VERSION : 0.1
   VAR_INPUT
      null_value : DInt;   // value that indicates null data
   END_VAR
   VAR_IN_OUT
      int_array : Variant;
   END_VAR
   VAR_TEMP
      i : Int;
      j : Int;
      len_int : Int;
      len_udint : UDInt;
      status : Int;
      t_int_array : Array[0..999] of DInt;
   END_VAR
BEGIN
   REGION "COPY TO LOCAL MEMORY"
       #len_udint := CountOfElements(#int_array);
       #len_int := UDINT_TO_INT(#len_udint) - 1;
       #status := MOVE_BLK_VARIANT(SRC := #int_array,
                                   COUNT := #len_udint,
                                   SRC_INDEX := 0,
                                   DEST_INDEX := 0,
                                   DEST => #t_int_array);
   END_REGION

   REGION "COLLAPSE IN PLACE"
       FOR #i := 0 TO #len_int - 1 DO
           IF #t_int_array[#i] = #null_value THEN
               FOR #j := #i + 1 TO #len_int DO
                   IF #t_int_array[#j] <> #null_value THEN
                       #t_int_array[#i] := #t_int_array[#j];
                       #t_int_array[#j] := #null_value;
                       EXIT;
                   END_IF;
               END_FOR;
           END_IF;
       END_FOR;
   END_REGION

   REGION "RETURN"
       #status := MOVE_BLK_VARIANT(SRC := #t_int_array,
                                   COUNT := #len_udint,
                                   SRC_INDEX := 0,
                                   DEST_INDEX := 0,
                                   DEST => #int_array);
   END_REGION
END_FUNCTION

FUNCTION "Count Collapsed DInt Array" : Int   // FC133, SCL
{ S7_Optimized_Access := 'TRUE' }
VERSION : 0.1
   VAR_INPUT
      null_value : DInt;
      "array" : Variant;
   END_VAR
   VAR_TEMP
      count : Int;
      i : Int;
      len_int : Int;
      len_udint : UDInt;
      status : Int;
      t_array : Array[0..999] of DInt;
   END_VAR
BEGIN
   REGION "NOTES"
       (*
       returns the number of valid elements in a collapsed int array
       *)
   END_REGION


   REGION "COPY TO LOCAL"
       #len_udint := CountOfElements(#array);
       #len_int := UDINT_TO_INT(#len_udint) - 1;
       #status := MOVE_BLK_VARIANT(SRC := #array,
                                   COUNT := #len_udint,
                                   SRC_INDEX := 0,
                                   DEST_INDEX := 0,
                                   DEST => #t_array);
   END_REGION


   REGION "SCAN FOR FIRST NULL"
       FOR #i := 0 TO #len_int DO
           IF #t_array[#i] = INT_TO_DINT("NULL_TOKEN") THEN
               EXIT;
           END_IF;
           IF #t_array[#i] <> #null_value THEN
               #count += 1;
           END_IF;
       END_FOR;
   END_REGION


   REGION "RETURN"
       #"Count Collapsed DInt Array" := #count;
   END_REGION
END_FUNCTION

FUNCTION "Map WIP Codes to DInt Array" : Void   // FC139, SCL
{ S7_Optimized_Access := 'TRUE' }
VERSION : 0.1
   VAR_INPUT
      station : "WIP: Station";
   END_VAR
   VAR_IN_OUT
      WIP_array : Array[0.."WIP_COUNT"] of DInt;
   END_VAR
   VAR_TEMP
      i : Int;
   END_VAR
BEGIN
   FOR #i := 0 TO "WIP_COUNT" DO
       IF #station.wip[#i].wip.code = "NULL_TOKEN" THEN
           EXIT;
       END_IF;
       #WIP_array[#i] := #station.wip[#i].wip.code;
   END_FOR;
END_FUNCTION

FUNCTION "Map Selected Stations to Int Array" : Void   // FC142, SCL
{ S7_Optimized_Access := 'TRUE' }
VERSION : 0.1
   VAR_INPUT
      selected_stations : "Selected Stations";
   END_VAR
   VAR_OUTPUT
      selected_stations_indicies : Array[0.."STATION_COUNT"] of Int;
   END_VAR
   VAR_TEMP
      i : Int;
      p_ret : Int;
      _return : Array[0.."STATION_COUNT"] of Int;
   END_VAR
BEGIN
   "Array.Int.Fill"(value := "NULL_TOKEN",
                    int_array := #_return);
   FOR #i := 0 TO "STATION_COUNT" DO
       IF #selected_stations.stns[#i] THEN
           #_return[#p_ret] := #i;
           #p_ret += 1;
       END_IF;
   END_FOR;
   #selected_stations_indicies := #_return;
END_FUNCTION

FUNCTION "Part_Number_Double.USInt_State_Change" : "State Changes: USInt"   // FC258, SCL
{ S7_Optimized_Access := 'TRUE' }
VERSION : 0.1
   VAR_INPUT
      interface : USInt;
      old : USInt;
   END_VAR
   VAR_TEMP
      _return : "State Changes: USInt";
   END_VAR
BEGIN
       #_return.rising := "USInt.Value_Change"(value := #interface,
                                               old_value := #old);
       #_return.actual := #interface;
       #_return.falling := FALSE;     // animate never set to null token 
       #"Part_Number_Double.USInt_State_Change" := #_return;
END_FUNCTION

FUNCTION "Part_Number_Double.Bool_State_Change" : "State Changes: Bool"   // FC259, SCL
{ S7_Optimized_Access := 'TRUE' }
VERSION : 0.1
   VAR_INPUT
      interface : Bool;
      old : Bool;
   END_VAR
   VAR_TEMP
      _return : "State Changes: Bool";
   END_VAR
BEGIN
   #_return.rising := "Bool.Rising_Edge"(signal := #interface,
                                                 old_signal := #old);
   #_return.actual := #interface;
   #_return.falling := "Bool.Falling_Edge"(signal := #interface,
                                           old_signal := #old);
   #"Part_Number_Double.Bool_State_Change" := #_return;
END_FUNCTION

FUNCTION "Part_Number_Double.WString_State_Change" : "State Changes: WString"   // FC260, SCL
{ S7_Optimized_Access := 'TRUE' }
VERSION : 0.1
   VAR_INPUT
      interface : WString;
      old : WString;
   END_VAR
   VAR_TEMP
      _return : "State Changes: WString";
   END_VAR
BEGIN
   #_return.rising := "WString.Rising_Edge"(value := #interface,
                                             old_value := #old);
   #_return.actual := #interface;
   #_return.falling := "WString.Falling_Edge"(value := #interface,
                                               old_value := #old);
   #"Part_Number_Double.WString_State_Change" := #_return;
END_FUNCTION

FUNCTION "Part_Number_Double_IO_Field.Set_Mode" : Void   // FC261, SCL
{ S7_Optimized_Access := 'TRUE' }
VERSION : 0.1
   VAR_INPUT
      feedback : "Part_Number_Double.State_Change.UDT";
   END_VAR
   VAR_IN_OUT
      mode : String;
   END_VAR
   VAR CONSTANT
      SINGLE : String := 'single';
      DOUBLE : String := 'double';
   END_VAR
BEGIN
   IF #mode = #SINGLE AND #feedback.single.actuate.falling THEN
       #mode := #DOUBLE;
       RETURN;
   END_IF;

   IF #mode = #DOUBLE AND #feedback.double.actuate.falling THEN
       #mode := #SINGLE;
       RETURN;
   END_IF;
END_FUNCTION

FUNCTION "Array.Table_Row.Copy" : Void   // FC296, SCL
{ S7_Optimized_Access := 'TRUE' }
VERSION : 0.1
   VAR_INPUT
      source : Array[*] of "Table Row";
   END_VAR
   VAR_IN_OUT
      destination : Array[*] of "Table Row";
   END_VAR
   VAR_TEMP
      _length_source : DInt;
      _length_destination : DInt;
      _upper_bound : DInt;
      _i : DInt;
   END_VAR
BEGIN
   REGION "FIND UPPER BOUND"
       #_length_source := UDINT_TO_DINT("Array.Any.Length"(#source)) - 1;
       #_length_destination := UDINT_TO_DINT("Array.Any.Length"(#destination)) - 1;
       #_upper_bound := #_length_source;
       IF #_length_destination < #_length_source THEN
           #_upper_bound := #_length_destination;
       END_IF;
   END_REGION


   REGION "PERFORM COPY"
       FOR #_i := 0 TO #_upper_bound DO
           #destination[#_i] := #source[#_i];
       END_FOR;
   END_REGION


   REGION "RETURN"    
       RETURN;
   END_REGION
END_FUNCTION

// folder: Utilities/Address

FUNCTION "Address.Get_Button" : DInt   // FC21, SCL
{ S7_Optimized_Access := 'TRUE' }
VERSION : 0.1
   VAR_INPUT
      address : DInt;
   END_VAR
BEGIN
   #"Address.Get_Button" := #address MOD 10;
END_FUNCTION

FUNCTION "Address.Get_Station" : DInt   // FC24, SCL
{ S7_Optimized_Access := 'TRUE' }
VERSION : 0.1
   VAR_INPUT
      address : DInt;
   END_VAR
BEGIN
   #"Address.Get_Station" := #address / 10_000;
END_FUNCTION

FUNCTION "Address.Set_Address" : DInt   // FC32, SCL
{ S7_Optimized_Access := 'TRUE' }
VERSION : 0.1
   VAR_INPUT
      pBtn : Int;
      pStn : Int;
      pWip : Int;
   END_VAR
BEGIN
   #"Address.Set_Address" := INT_TO_DINT(#pStn) * 10_000 + INT_TO_DINT(#pWip) * 10 + INT_TO_DINT(#pBtn);
END_FUNCTION

FUNCTION "Address.Get_Wip" : DInt   // FC88, SCL
{ S7_Optimized_Access := 'TRUE' }
VERSION : 0.1
   VAR_INPUT
      address : DInt;
   END_VAR
BEGIN
   #"Address.Get_Wip" := #address - "Address.Get_Station"(#address) * 10_000 - "Address.Get_Button"(#address);
END_FUNCTION

// folder: Utilities/Array

FUNCTION "Array.Any.Length" : UDInt   // FC60, SCL
{ S7_Optimized_Access := 'TRUE' }
VERSION : 0.1
   VAR_INPUT
      "array" : Variant;
   END_VAR
   VAR_TEMP
      status : DInt;
      ret : UDInt;
   END_VAR
BEGIN
   #ret := CountOfElements(#array);
   #"Array.Any.Length" := #ret;
END_FUNCTION

FUNCTION "Get Station Index From Id" : Int   // FC106, SCL
{ S7_Optimized_Access := 'TRUE' }
VERSION : 0.1
   VAR_INPUT
      line_name : WString;
      drop_zone : USInt;
      stns : "Station: All Stations";
   END_VAR
   VAR_TEMP
      i : Int;
      ret : Int;
   END_VAR
BEGIN
   REGION "MATCH LINE NAME AND DROP ZONE"
       FOR #i := 0 TO "STATION_COUNT" DO
           IF #line_name = #stns.stn[#i].id.lineName THEN
               IF #drop_zone = #stns.stn[#i].id.dropZone THEN
                   #ret := #i;
                   EXIT;
               END_IF;
           END_IF;
       END_FOR;
   END_REGION


   REGION "RETURN"
       #"Get Station Index From Id" := #ret;
   END_REGION
END_FUNCTION

FUNCTION "Array.Int.Fill" : Void   // FC109, SCL
{ S7_Optimized_Access := 'TRUE' }
VERSION : 0.1
   VAR_INPUT
      value : Int;
   END_VAR
   VAR_IN_OUT
      int_array : Array[*] of Int;
   END_VAR
   VAR_TEMP
      _i : DInt;
      _length : DInt;
   END_VAR
BEGIN
   REGION "GET LENGHT"
       #_length := UDINT_TO_DINT("Array.Any.Length"(#int_array));
       #_length -= 1;
   END_REGION


   REGION "FILL LENGTH WITH BYTE IN"
       FOR #_i := 0 TO #_length DO
           #int_array[#_i] := #value;
       END_FOR;
   END_REGION
END_FUNCTION

FUNCTION "Array.DInt.Is_Element" : Bool   // FC111, SCL
{ S7_Optimized_Access := 'TRUE' }
VERSION : 0.1
   VAR_INPUT
      dint_array : Array[*] of DInt;
      search_term : DInt;
   END_VAR
   VAR_TEMP
      _i : DInt;
      _length : DInt;
   END_VAR
BEGIN
   REGION "LOCAL VARIABLES"
       #_length := UDINT_TO_DINT("Array.Any.Length"(#dint_array)) - 1;
   END_REGION


   REGION "SEARCH ARRAY"
       FOR #_i := 0 TO #_length DO
           IF #dint_array[#_i] <> #search_term THEN
               CONTINUE;
           END_IF;
           #"Array.DInt.Is_Element" := TRUE;
           RETURN;
       END_FOR;
   END_REGION


   REGION "NOT FOUND"
       #"Array.DInt.Is_Element" := FALSE;
       RETURN;
   END_REGION
END_FUNCTION

FUNCTION "Array.Int.Collapse" : Void   // FC114, SCL
{ S7_Optimized_Access := 'TRUE' }
VERSION : 0.1
   VAR_INPUT
      null_value : Int;   // value that indicates null data
   END_VAR
   VAR_IN_OUT
      int_array : Variant;
   END_VAR
   VAR_TEMP
      i : Int;
      j : Int;
      len_int : Int;
      len_udint : UDInt;
      status : Int;
      t_int_array : Array[0..999] of Int;
   END_VAR
BEGIN
   REGION "COPY TO LOCAL MEMORY"
       #len_udint := CountOfElements(#int_array);
       #len_int := UDINT_TO_INT(#len_udint) - 1;
       #status := MOVE_BLK_VARIANT(SRC := #int_array,
                                   COUNT := #len_udint,
                                   SRC_INDEX := 0,
                                   DEST_INDEX := 0,
                                   DEST => #t_int_array);
   END_REGION

   REGION "COLLAPSE IN PLACE"
       FOR #i := 0 TO #len_int - 1 DO
           IF #t_int_array[#i] = #null_value THEN
               FOR #j := #i + 1 TO #len_int DO
                   IF #t_int_array[#j] <> #null_value THEN
                       #t_int_array[#i] := #t_int_array[#j];
                       #t_int_array[#j] := #null_value;
                       EXIT;
                   END_IF;
               END_FOR;
           END_IF;
       END_FOR;
   END_REGION

   REGION "RETURN"
       #status := MOVE_BLK_VARIANT(SRC := #t_int_array,
                                   COUNT := #len_udint,
                                   SRC_INDEX := 0,
                                   DEST_INDEX := 0,
                                   DEST => #int_array);
   END_REGION
END_FUNCTION

FUNCTION "Array.Int.Count" : Int   // FC115, SCL
{ S7_Optimized_Access := 'TRUE' }
VERSION : 0.1
   VAR_INPUT
      null_value : Int;
      "array" : Variant;
   END_VAR
   VAR_TEMP
      count : Int;
      i : Int;
      len_int : Int;
      len_udint : UDInt;
      status : Int;
      t_array : Array[0..999] of Int;
   END_VAR
BEGIN
   REGION "NOTES"
       (*
       returns the number of valid elements in a collapsed int array
       *)
   END_REGION


   REGION "COPY TO LOCAL"
       #len_udint := CountOfElements(#array);
       #len_int := UDINT_TO_INT(#len_udint) - 1;
       #status := MOVE_BLK_VARIANT(SRC := #array,
                                   COUNT := #len_udint,
                                   SRC_INDEX := 0,
                                   DEST_INDEX := 0,
                                   DEST => #t_array);
   END_REGION


   REGION "SCAN FOR FIRST NULL"
       FOR #i := 0 TO #len_int DO
           IF #t_array[#i] = #null_value THEN
               EXIT;
           END_IF;
           IF #t_array[#i] <> #null_value THEN
               #count += 1;
           END_IF;
       END_FOR;
   END_REGION


   REGION "RETURN"
       #"Array.Int.Count" := #count;
   END_REGION
END_FUNCTION

FUNCTION "Array.Bool.True_Indices" : Void   // FC120, SCL
{ S7_Optimized_Access := 'TRUE' }
VERSION : 0.1
   VAR_INPUT
      array_of_bool : Array[*] of Bool;   // max 1000 elements
      length : Int;   // necessary because dynamically sized arrays of bool get passed as arrays with size of a multiple of 8
   END_VAR
   VAR_IN_OUT
      list_of_indices : Array[*] of Int;   // max 1000 elements
   END_VAR
   VAR_TEMP
      _i : Int;
      _p_return : Int;
      _resized_bool_array : Array[0..#UBOUND] of Bool;
   END_VAR
   VAR CONSTANT
      UBOUND : Int := 999;
   END_VAR
BEGIN
   REGION "FILL RETURN ARRAY"
       "Array.Int.Fill"(value := "NULL_TOKEN",
                        int_array := #list_of_indices);
   END_REGION


   REGION "COPY TO ARRAY OF STATIC SIZE"
       FOR #_i := 0 TO #length DO
           #_resized_bool_array[#_i] := #array_of_bool[#_i];
       END_FOR;
   END_REGION


   REGION "INSERT INDICES INTO RETURN ARRAY"
       FOR #_i := 0 TO #length DO
           IF #_resized_bool_array[#_i] THEN
               #list_of_indices[#_p_return] := #_i;
               #_p_return += 1;
           END_IF;
       END_FOR;
   END_REGION
END_FUNCTION

FUNCTION "Array.Int.Is_Element" : Bool   // FC121, SCL
{ S7_Optimized_Access := 'TRUE' }
VERSION : 0.1
   VAR_INPUT
      int_array : Array[*] of Int;
      search_term : Int;
   END_VAR
   VAR_TEMP
      _i : Int;
      _length : DInt;
   END_VAR
BEGIN
   REGION "LOCAL VARIABLES"
       #_length := UDINT_TO_DINT("Array.Any.Length"(#int_array)) - 1;
   END_REGION


   REGION "SEARCH ARRAY"
       FOR #_i := 0 TO #_length DO
           IF #int_array[#_i] <> #search_term THEN
               CONTINUE;
           END_IF;
           #"Array.Int.Is_Element" := TRUE;
           RETURN;
       END_FOR;
   END_REGION


   REGION "NOT FOUND"
       #"Array.Int.Is_Element" := FALSE;
       RETURN;
   END_REGION
END_FUNCTION

FUNCTION "Array.DInt.Fill" : Void   // FC131, SCL
{ S7_Optimized_Access := 'TRUE' }
VERSION : 0.1
   VAR_INPUT
      int_in : DInt;
   END_VAR
   VAR_OUTPUT
      array_out : Variant;
   END_VAR
   VAR_TEMP
      i : Int;
      internal_array : Array[0..999] of DInt;
      len_array_out : UDInt;
      status : Int;
   END_VAR
BEGIN
   REGION "GET LENGHT"
       #len_array_out := CountOfElements(#array_out);
   END_REGION


   REGION "FILL LENGTH WITH BYTE IN"
       FOR #i := 0 TO UDINT_TO_INT(#len_array_out) - 1 DO
           #internal_array[#i] := #int_in;
       END_FOR;
   END_REGION


   REGION "RETURN"
       #status := MOVE_BLK_VARIANT(SRC := #internal_array,
                                   COUNT := #len_array_out,
                                   SRC_INDEX := 0,
                                   DEST_INDEX := 0,
                                   DEST => #array_out);
   END_REGION
END_FUNCTION

FUNCTION "Array.Int.Search" : Int   // FC140, SCL
{ S7_Optimized_Access := 'TRUE' }
VERSION : 0.1
   VAR_INPUT
      array_of_int : Variant;   // max upper bound 999
      search_term : Int;
   END_VAR
   VAR_TEMP
      i : Int;
      len_as_udint : UDInt;
      len_as_int : Int;
      ret : Int;
      status : Int;
      t_array : Array[0..999] of Int;
   END_VAR
   // Ret_Val : index of search term. returns -1 if not found.
BEGIN
   REGION "LOCAL VARIABLES"
       #len_as_udint := CountOfElements(#array_of_int);
       #len_as_int := UDINT_TO_INT(#len_as_udint) - 1;
       #status := MOVE_BLK_VARIANT(SRC := #array_of_int,
                                   COUNT := #len_as_udint,
                                   SRC_INDEX := 0,
                                   DEST_INDEX := 0,
                                   DEST => #t_array);
       #ret := -1;
   END_REGION


   REGION "SEARCH ARRAY"
       FOR #i := 0 TO #len_as_int DO
           IF #t_array[#i] = #search_term THEN
               #ret := #i;
               EXIT;
           END_IF;
       END_FOR;
   END_REGION


   REGION "RETURN"
       #"Array.Int.Search" := #ret;
   END_REGION
END_FUNCTION

FUNCTION "Array.Int.Intersect" : Void   // FC141, SCL
{ S7_Optimized_Access := 'TRUE' }
VERSION : 0.1
   VAR_INPUT
      "a" : Variant;   // should be array of int, max 999
      "b" : Variant;   // should be array of int, max 999
      null_value : Int;
   END_VAR
   VAR_OUTPUT
      intersect_array : Variant;   // should be array of int, max 999
   END_VAR
   VAR_TEMP
      i : Int;
      j : Int;
      len_a : Struct
         as_udint : UDInt;
         as_int : Int;
      END_STRUCT;
      len_b : Struct
         as_udint : UDInt;
         as_int : Int;
      END_STRUCT;
      len_longer : Struct
         as_udint : UDInt;
         as_int : Int;
      END_STRUCT;
      len_shorter : Struct
         as_udint : UDInt;
         as_int : Int;
      END_STRUCT;
      t_a : Array[0..#u_bound] of Int;
      p_ret : Int;
      ret : Array[0..#u_bound_double] of Int;
      t_b : Array[0..#u_bound] of Int;
      status : Int;
   END_VAR
   VAR CONSTANT
      u_bound : Int := 999;
      u_bound_double : Int := 1999;
   END_VAR
BEGIN
   REGION "GET LENGTHS"
       #len_a.as_udint := CountOfElements(#a);
       #len_a.as_int := UDINT_TO_INT(#len_a.as_udint) - 1;
       #len_b.as_udint := CountOfElements(#b);
       #len_b.as_int := UDINT_TO_INT(#len_b.as_udint) - 1;
   END_REGION

   REGION "MOVE"
       #status := MOVE_BLK_VARIANT(SRC := #a, COUNT := #len_a.as_udint, SRC_INDEX := 0, DEST_INDEX := 0, DEST => #t_a);
       #status := MOVE_BLK_VARIANT(SRC := #b, COUNT := #len_b.as_udint, SRC_INDEX := 0, DEST_INDEX := 0, DEST => #t_b);
   END_REGION

   REGION "FIND INTERSECT"
       FOR #i := 0 TO #len_a.as_int DO
           IF #t_a[#i] = #null_value THEN
               EXIT;
           END_IF;
           FOR #j := 0 TO #len_b.as_int DO
               IF #t_b[#j] = #null_value THEN
                   EXIT;
               END_IF;
               IF #t_a[#i] = #t_b[#j] THEN
                   #ret[#p_ret] := #t_a[#i];
                   #p_ret += 1;
                   EXIT;
               END_IF;
           END_FOR;
       END_FOR;
   END_REGION

   REGION "RETURN"
       #status := MOVE_BLK_VARIANT(SRC := #ret, COUNT := INT_TO_UDINT(#p_ret - 1), SRC_INDEX := 0, DEST_INDEX := 0, DEST => #intersect_array);
   END_REGION
END_FUNCTION

FUNCTION "Array.DInt.First_Occurance" : DInt   // FC143, SCL
{ S7_Optimized_Access := 'TRUE' }
VERSION : 0.1
   VAR_INPUT
      dint_array : Array[*] of DInt;
      search_term : Int;
   END_VAR
   VAR_TEMP
      _i : DInt;
      _length : UDInt;
   END_VAR
BEGIN
   REGION "NOTES"
       (* 
       This function returns the first occurance of the search term.
       This function meant for use with collapsed arrays.
       See "Array.DInt.Collapse" for collapse functionality.
       *)
   END_REGION


   REGION "GET LENGTH OF INPUT ARRAY"
       #_length := "Array.Any.Length"(#dint_array);
   END_REGION


   REGION "FIND FIRST SEARCH TERM, -1 IF NONE"
       (*
       Its worth noting that "Array.DInt.Is_Element" could return the index of the search term
       as an output, saving the processor some work. 
       The rework is justified by increased encapsulation.
       The time complexity for "Array.DInt.First_Occurance" remains O(n).
       *)
       IF NOT "Array.DInt.Is_Element"(dint_array := #dint_array, search_term := #search_term) THEN
           #"Array.DInt.First_Occurance" := -1;
           RETURN;
       END_IF;
       WHILE #dint_array[#_i] <> #search_term AND DINT_TO_UDINT(#_i) < #_length DO
           #_i += 1;
       END_WHILE;
   END_REGION


   REGION _name_
       #"Array.DInt.First_Occurance" := #_i;
   END_REGION
END_FUNCTION

FUNCTION "Array.DInt.Intersect_Exists" : Bool   // FC144, SCL
{ S7_Optimized_Access := 'TRUE' }
VERSION : 0.1
   VAR_INPUT
      "a" : Variant;   // should be array of dint, max 999
      "b" : Variant;   // should be array of dint, max 999
      null_value : DInt;
   END_VAR
   VAR_TEMP
      i : Int;
      j : Int;
      len_a : Struct
         as_udint : UDInt;
         as_int : Int;
      END_STRUCT;
      len_b : Struct
         as_udint : UDInt;
         as_int : Int;
      END_STRUCT;
      t_a : Array[0..#u_bound] of DInt;
      p_ret : Int;
      ret : Bool;
      t_b : Array[0..#u_bound] of DInt;
      status : Int;
   END_VAR
   VAR CONSTANT
      u_bound : Int := 999;
   END_VAR
BEGIN
   REGION "GET LENGHTS"
       #len_a.as_udint := CountOfElements(#a);
       #len_a.as_int := UDINT_TO_INT(#len_a.as_udint) - 1;
       #len_b.as_udint := CountOfElements(#b);
       #len_b.as_int := UDINT_TO_INT(#len_b.as_udint) - 1;
   END_REGION

   REGION "PERFORM MOVES"
       #status := MOVE_BLK_VARIANT(SRC := #a, COUNT := #len_a.as_udint, SRC_INDEX := 0, DEST_INDEX := 0, DEST => #t_a);
       #status := MOVE_BLK_VARIANT(SRC := #b, COUNT := #len_b.as_udint, SRC_INDEX := 0, DEST_INDEX := 0, DEST => #t_b);
   END_REGION


   REGION "SEARCH FOR ANY MATCHING ELEMENT"
       FOR #i := 0 TO #len_a.as_int DO

           REGION "SKIP NULL VALUES"
               IF #t_a[#i] = #null_value THEN
                   CONTINUE;
               END_IF;
           END_REGION

           REGION "INNER LOOP"
               FOR #j := 0 TO #len_b.as_int DO

                   REGION "SKIP NULL VALUES"
                       IF #t_b[#j] = #null_value THEN
                           CONTINUE;
                       END_IF;
                   END_REGION

                   REGION "SET RETURN VALUE ON MATCH"
                       IF #t_a[#i] = #t_b[#j] THEN
                           #ret := TRUE;
                           EXIT;
                       END_IF;
                   END_REGION

               END_FOR;
           END_REGION

           REGION "EXIT OUTTER LOOP IF MATCH FOUND"
               IF #ret THEN
                   EXIT;
               END_IF;
           END_REGION

       END_FOR;
   END_REGION

   REGION "RETURN"
       #"Array.DInt.Intersect_Exists" := #ret;
   END_REGION
END_FUNCTION

FUNCTION "Array.DInt.Intersect" : Void   // FC145, SCL
{ S7_Optimized_Access := 'TRUE' }
VERSION : 0.1
   VAR_INPUT
      "a" : Variant;   // should be array of dint, max 999
      "b" : Variant;   // should be array of dint, max 999
      null_value : DInt;
   END_VAR
   VAR_OUTPUT
      intersect_array : Variant;   // should be array of dint, max 999
   END_VAR
   VAR_TEMP
      i : Int;
      j : Int;
      len_a : Struct
         as_udint : UDInt;
         as_int : Int;
      END_STRUCT;
      len_b : Struct
         as_udint : UDInt;
         as_int : Int;
      END_STRUCT;
      t_a : Array[0..#u_bound] of DInt;
      p_ret : Int;
      ret : Array[0..#u_bound_double] of DInt;
      t_b : Array[0..#u_bound] of DInt;
      status : Int;
   END_VAR
   VAR CONSTANT
      u_bound : Int := 999;
      u_bound_double : Int := 1999;
   END_VAR
BEGIN
   REGION "GET LENGTHS"
       #len_a.as_udint := CountOfElements(#a);
       #len_a.as_int := UDINT_TO_INT(#len_a.as_udint) - 1;
       #len_b.as_udint := CountOfElements(#b);
       #len_b.as_int := UDINT_TO_INT(#len_b.as_udint) - 1;
   END_REGION

   REGION "MOVE"
       #status := MOVE_BLK_VARIANT(SRC := #a, COUNT := #len_a.as_udint, SRC_INDEX := 0, DEST_INDEX := 0, DEST => #t_a);
       #status := MOVE_BLK_VARIANT(SRC := #b, COUNT := #len_b.as_udint, SRC_INDEX := 0, DEST_INDEX := 0, DEST => #t_b);
   END_REGION

   REGION "FIND INTERSECT"
       FOR #i := 0 TO #len_a.as_int DO
           IF #t_a[#i] = #null_value THEN
               EXIT;
           END_IF;
           FOR #j := 0 TO #len_b.as_int DO
               IF #t_b[#j] = #null_value THEN
                   EXIT;
               END_IF;
               IF #t_a[#i] = #t_b[#j] THEN
                   #ret[#p_ret] := #t_a[#i];
                   #p_ret += 1;
                   EXIT;
               END_IF;
           END_FOR;
       END_FOR;
   END_REGION

   REGION "RETURN"
       #status := MOVE_BLK_VARIANT(SRC := #ret, COUNT := INT_TO_UDINT(#p_ret - 1), SRC_INDEX := 0, DEST_INDEX := 0, DEST => #intersect_array);
   END_REGION
END_FUNCTION

FUNCTION "Array.WString.Is_Element" : Bool   // FC207, SCL
{ S7_Optimized_Access := 'TRUE' }
VERSION : 0.1
   VAR_INPUT
      search_term : WString;
      search_array : Array[*] of WString[1];
   END_VAR
   VAR_TEMP
      _i : Int;
      _length_search_array : UDInt;
   END_VAR
BEGIN
   #_length_search_array := "Array.Any.Length"(#search_array);
   FOR #_i := 0 TO UDINT_TO_INT(#_length_search_array - 1) DO
       IF #search_term = #search_array[#_i] THEN
           #"Array.WString.Is_Element" := TRUE;
           RETURN;
       END_IF;
   END_FOR;
   #"Array.WString.Is_Element" := FALSE;
END_FUNCTION

FUNCTION "Array.Int.First_Occurance" : DInt   // FC220, SCL
{ S7_Optimized_Access := 'TRUE' }
VERSION : 0.1
   VAR_INPUT
      int_array : Array[*] of Int;
      search_term : Int;
   END_VAR
   VAR_TEMP
      _i : DInt;
      _length : UDInt;
   END_VAR
BEGIN
   REGION "NOTES"
       (* 
       This function returns the first occurance of the search term.
       This function meant for use with collapsed arrays.
       See "Array.Int.Collapse" for collapse functionality.
       *)
   END_REGION


   REGION "GET LENGTH OF INPUT ARRAY"
       #_length := "Array.Any.Length"(#int_array);
   END_REGION


   REGION "FIND FIRST SEARCH TERM, -1 IF NONE"
       (*
       Its worth noting that "Array.Int.Is_Element" could return the index of the search term
       as an output, saving the processor some work. 
       The rework is justified by increased encapsulation.
       The time complexity for "Array.Int.First_Occurance" remains O(n).
       *)
       IF NOT "Array.Int.Is_Element"(int_array := #int_array, search_term := #search_term) THEN
           #"Array.Int.First_Occurance" := -1;
           RETURN;
       END_IF;
       WHILE #int_array[#_i] <> #search_term AND DINT_TO_UDINT(#_i) < #_length DO
           #_i += 1;
       END_WHILE;
   END_REGION


   REGION _name_
       #"Array.Int.First_Occurance" := #_i;
   END_REGION
END_FUNCTION

FUNCTION "Array.WString.Fill" : Void   // FC243, SCL
{ S7_Optimized_Access := 'TRUE' }
VERSION : 0.1
   VAR_INPUT
      value : WString;
   END_VAR
   VAR_IN_OUT
      "array" : Array[*] of WString;
   END_VAR
   VAR_TEMP
      _length : Int;
      _i : Int;
   END_VAR
BEGIN
   #_length := UDINT_TO_INT("Array.Any.Length"(#array)) - 1;
   FOR #_i := 0 TO #_length DO
       #array[#_i] := #value;
   END_FOR;
   RETURN;
END_FUNCTION

FUNCTION "Array.WString.Search" : Int   // FC244, SCL
{ S7_Optimized_Access := 'TRUE' }
VERSION : 0.1
   VAR_INPUT
      "array" : Array[*] of WString;
      search_term : WString;
   END_VAR
   VAR_TEMP
      _i : Int;
      _length : Int;
   END_VAR
   // Ret_Val : index of search term. returns -1 if not found.
BEGIN
   REGION "SEARCH ARRAY"    
       #_length := UDINT_TO_INT("Array.Any.Length"(#array)) - 1;
       FOR #_i := 0 TO #_length DO
           IF #array[#_i] = #search_term THEN
               #"Array.WString.Search" := #_i;
               RETURN;
           END_IF;
       END_FOR;
   END_REGION

   REGION "RETURN"
       #"Array.WString.Search" := "NULL_TOKEN";
       RETURN;
   END_REGION
END_FUNCTION

FUNCTION "Array.Char.Search" : Int   // FC266, SCL
{ S7_Optimized_Access := 'TRUE' }
VERSION : 0.1
   VAR_INPUT
      "array" : Array[*] of Char;   // max upper bound 999
      search_term : Char;
   END_VAR
   VAR_TEMP
      _i : Int;
      _length : Int;
   END_VAR
   // Ret_Val : index of search term. returns -1 if not found.
BEGIN
   REGION "GET LENGTH"
       #_length := UDINT_TO_INT("Array.Any.Length"(#array)) - 1;
   END_REGION


   REGION "SEARCH ARRAY"
       FOR #_i := 0 TO #_length DO
           IF #array[#_i] = #search_term THEN
               #"Array.Char.Search" := #_i;
               EXIT;
           END_IF;
       END_FOR;
   END_REGION


   REGION "RETURN"
       #"Array.Char.Search" := "NULL_TOKEN";
   END_REGION
END_FUNCTION

FUNCTION "Array.WString.Reverse" : Void   // FC270, SCL
{ S7_Optimized_Access := 'TRUE' }
VERSION : 0.1
   VAR_INPUT
      null_token : WString;
   END_VAR
   VAR_IN_OUT
      wstring_array : Array[*] of WString;
   END_VAR
   VAR_TEMP
      _has_data_count : Int;
      _i : Int;
      _p_swap : Int;
      _temp : WString;
   END_VAR
   VAR CONSTANT
      NOT_FOUND : Int := -1;
   END_VAR
BEGIN
   REGION "CHECK FOR FIRST EMPTY POSITION"
       #_has_data_count := "Array.WString.Search"(array := #wstring_array,
                                                  search_term := #null_token);
   END_REGION


   REGION "EXIT ON EMPTY ARRAY"
       IF #_has_data_count = 0 THEN
           RETURN;
       END_IF;
   END_REGION


   REGION "ARRAY IS FULL"
       IF #_has_data_count = #NOT_FOUND THEN
           #_has_data_count := UDINT_TO_INT("Array.Any.Length"(#wstring_array));
       END_IF;
   END_REGION


   REGION "ADJUST TO ZERO INDEX"
       #_has_data_count -= 1;
   END_REGION


   REGION "SWAP ELEMENTS"
       FOR #_i := 0 TO #_has_data_count / 2 DO
           #_p_swap := #_has_data_count - #_i;
           #_temp := #wstring_array[#_i];
           #wstring_array[#_i] := #wstring_array[#_p_swap];
           #wstring_array[#_p_swap] := #_temp;
       END_FOR;
   END_REGION


   REGION "DONE"
       RETURN;
   END_REGION
END_FUNCTION

FUNCTION "Array.DInt.Search" : DInt   // FC305, SCL
{ S7_Optimized_Access := 'TRUE' }
VERSION : 0.1
   VAR_INPUT
      array_of_int : Variant;   // max upper bound 999
      search_term : DInt;
   END_VAR
   VAR_TEMP
      _i : Int;
      _len_as_udint : UDInt;
      _len_as_int : Int;
      _status : Int;
      _t_array : Array[0..999] of Int;
   END_VAR
   // Ret_Val : index of search term. returns -1 if not found.
BEGIN
   REGION "LOCAL VARIABLES"
       #_len_as_udint := CountOfElements(#array_of_int);
       #_len_as_int := UDINT_TO_INT(#_len_as_udint) - 1;
       #_status := MOVE_BLK_VARIANT(SRC := #array_of_int,
                                    COUNT := #_len_as_udint,
                                    SRC_INDEX := 0,
                                    DEST_INDEX := 0,
                                    DEST => #_t_array);
   END_REGION


   REGION "SEARCH ARRAY"
       FOR #_i := 0 TO #_len_as_int DO
           IF #_t_array[#_i] <> #search_term THEN
               CONTINUE;
           END_IF;
           #"Array.DInt.Search" := #_i;
           RETURN;
       END_FOR;
   END_REGION


   REGION "RETURN"
       #"Array.DInt.Search" := INT_TO_DINT("NULL_TOKEN");
       RETURN;
   END_REGION
END_FUNCTION

// folder: Utilities/Bool

FUNCTION "Bool.Animate" : USInt   // FC9, SCL
{ S7_Optimized_Access := 'TRUE' }
VERSION : 0.1
   VAR_INPUT
      true_color : USInt;
      false_color : USInt;
      evaluation_signal : Bool;
   END_VAR
   VAR_TEMP
      animate : USInt;
   END_VAR
BEGIN
   REGION "FALSE COLOR"
       IF NOT #evaluation_signal THEN
           #animate := #false_color;
       END_IF;
   END_REGION

   REGION "TRUE COLOR"
       IF #evaluation_signal THEN
           #animate := #true_color;
       END_IF;
   END_REGION

   REGION "FUNCTION RETURN"
       #"Bool.Animate" := #animate;
   END_REGION
END_FUNCTION

FUNCTION "Bool.Rising_Edge" : Bool   // FC177, SCL
{ S7_Optimized_Access := 'TRUE' }
VERSION : 0.1
   VAR_INPUT
      signal : Bool;
      old_signal : Bool;
   END_VAR
BEGIN
   #"Bool.Rising_Edge" := #signal AND NOT #old_signal;
END_FUNCTION

FUNCTION "Bool.Falling_Edge" : Bool   // FC178, SCL
{ S7_Optimized_Access := 'TRUE' }
VERSION : 0.1
   VAR_INPUT
      signal : Bool;
      old_signal : Bool;
   END_VAR
BEGIN
   #"Bool.Falling_Edge" := NOT #signal AND #old_signal;
END_FUNCTION

// folder: Utilities/DInt

FUNCTION "Pointer Calc: KP8 Labels" : Int   // FC25, SCL
{ S7_Optimized_Access := 'TRUE' }
VERSION : 0.1
   VAR_INPUT
      index : Int;
   END_VAR
   VAR_TEMP
      val : Int;
   END_VAR
BEGIN
   IF #index >= 4 THEN
       #val := 7 - (#index - 4) * 2;
   END_IF;

   IF #index <= 3 THEN
       #val := 8 - #index * 2;
   END_IF;

   #"Pointer Calc: KP8 Labels" := #val;
END_FUNCTION

FUNCTION "DInt.Clip.Maximum" : DInt   // FC224, SCL
{ S7_Optimized_Access := 'TRUE' }
VERSION : 0.1
   VAR_INPUT
      value : DInt;
      maximum : DInt;
   END_VAR
BEGIN
   IF #value > #maximum THEN
       #"DInt.Clip.Maximum" := #maximum;
       RETURN;
   END_IF;
   #"DInt.Clip.Maximum" := #value;
END_FUNCTION

FUNCTION "DInt.Clip.Minimum" : DInt   // FC225, SCL
{ S7_Optimized_Access := 'TRUE' }
VERSION : 0.1
   VAR_INPUT
      value : DInt;
      minimum : DInt;
   END_VAR
BEGIN
   IF #value < #minimum THEN
       #"DInt.Clip.Minimum" := #minimum;
       RETURN;
   END_IF;
   #"DInt.Clip.Minimum" := #value;
END_FUNCTION

FUNCTION "DInt.Clip.Range" : DInt   // FC227, SCL
{ S7_Optimized_Access := 'TRUE' }
VERSION : 0.1
   VAR_INPUT
      value : DInt;
      maximum : DInt;
      minimum : DInt;
   END_VAR
   VAR_TEMP
      _return : DInt;
   END_VAR
BEGIN
   #_return := #value;
   #_return := "DInt.Clip.Maximum"(value := #value, maximum := #minimum);
   #_return := "DInt.Clip.Minimum"(value := #value, minimum := #minimum);
   #"DInt.Clip.Range" := #_return;
END_FUNCTION

// folder: Utilities/Int

FUNCTION "Int.Value_Change" : Bool   // FC179, SCL
{ S7_Optimized_Access := 'TRUE' }
VERSION : 0.1
   VAR_INPUT
      value : Int;
      old_value : Int;
   END_VAR
BEGIN
   #"Int.Value_Change" := #value <> #old_value;
END_FUNCTION

FUNCTION "Int.Clip.Minimum" : Int   // FC222, SCL
{ S7_Optimized_Access := 'TRUE' }
VERSION : 0.1
   VAR_INPUT
      value : Int;
      minimum : Int;
   END_VAR
BEGIN
   IF #value < #minimum THEN
       #"Int.Clip.Minimum" := #minimum;
       RETURN;
   END_IF;
   #"Int.Clip.Minimum" := #value;
END_FUNCTION

FUNCTION "Int.Clip.Maximum" : Int   // FC223, SCL
{ S7_Optimized_Access := 'TRUE' }
VERSION : 0.1
   VAR_INPUT
      value : Int;
      maximum : Int;
   END_VAR
BEGIN
   IF #value > #maximum THEN
       #"Int.Clip.Maximum" := #maximum;
       RETURN;
   END_IF;
   #"Int.Clip.Maximum" := #value;
END_FUNCTION

FUNCTION "Int.Clip.Range" : Int   // FC226, SCL
{ S7_Optimized_Access := 'TRUE' }
VERSION : 0.1
   VAR_INPUT
      value : Int;
      maximum : Int;
      minimum : Int;
   END_VAR
   VAR_TEMP
      _return : Int;
   END_VAR
BEGIN
   #_return := #value;
   #_return := "Int.Clip.Maximum"(value := #_return, maximum := #maximum);
   #_return := "Int.Clip.Minimum"(value:=#_return, minimum:=#minimum);
   #"Int.Clip.Range" := #_return;
END_FUNCTION

// folder: Utilities/NavBar

FUNCTION_BLOCK "NavBar: Top"   // FB31, SCL
{ S7_Optimized_Access := 'TRUE' }
VERSION : 0.1
   VAR_INPUT
      hide : Bool;
      TABLE_LENGTH : DInt;
   END_VAR
   VAR_IN_OUT
      interface : "Push Button Data";
      first_row : DInt;
   END_VAR
   VAR
      "Get Button Feedback" : "Push Button: State Changes";
   END_VAR
   VAR_TEMP
      feedback : "Push Button Data: State Change Data";
   END_VAR
BEGIN
   REGION "PROCESS USER INPUT"
       #"Get Button Feedback"(interface := #interface,
                              state_changes := #feedback);
   END_REGION

   REGION "ANIMATIONS"

       REGION "COLOR"
           #interface.animate := "Bool.Animate"(true_color := "GREEN_LIGHT_BACKGROUND",
                                                false_color := "GRAY_BACKGROUND",
                                                evaluation_signal := #feedback.actuate.actual);
       END_REGION

       REGION "VISIBILITY"
           #interface.visible := NOT #hide;
       END_REGION

       REGION "ENABLED STATE"
           #interface.enable := NOT #hide;
       END_REGION

   END_REGION

   REGION "SET FIRST ROW"
       IF #feedback.actuate.rising THEN
           #first_row := 0;
       END_IF;
   END_REGION
END_FUNCTION_BLOCK

FUNCTION_BLOCK "NavBar: Bottom"   // FB32, SCL
{ S7_Optimized_Access := 'TRUE' }
VERSION : 0.1
   VAR_INPUT
      hide : Bool;
      TABLE_LENGTH : DInt;
      VISIBLE_ROW_COUNT : DInt;
   END_VAR
   VAR_IN_OUT
      interface : "Push Button Data";
      first_row : DInt;
   END_VAR
   VAR
      "Get Button Feedback" : "Push Button: State Changes";
   END_VAR
   VAR_TEMP
      feedback : "Push Button Data: State Change Data";
   END_VAR
BEGIN
   REGION "PROCESS USER INPUT"
       #"Get Button Feedback"(interface := #interface,
                              state_changes := #feedback);
   END_REGION

   REGION "ANIMATIONS"

       REGION "COLOR"
           #interface.animate := "Bool.Animate"(true_color := "GREEN_LIGHT_BACKGROUND",
                                                false_color := "GRAY_BACKGROUND",
                                                evaluation_signal := #feedback.actuate.actual);
       END_REGION

       REGION "VISIBILITY"
           #interface.visible := NOT #hide;
       END_REGION

       REGION "ENABLED STATE"
           #interface.enable := NOT #hide;
       END_REGION

   END_REGION


   REGION "SET FIRST ROW"
       IF #feedback.actuate.rising THEN
           #first_row := #TABLE_LENGTH - #VISIBLE_ROW_COUNT;
       END_IF;
   END_REGION
END_FUNCTION_BLOCK

FUNCTION_BLOCK "NavBar: Page Up"   // FB36, SCL
{ S7_Optimized_Access := 'TRUE' }
VERSION : 0.1
   VAR_INPUT
      hide : Bool;
      TABLE_LENGTH : DInt;
      VISIBLE_ROW_COUNT : DInt;
   END_VAR
   VAR_IN_OUT
      interface : "Push Button Data";
      first_row : DInt;
   END_VAR
   VAR
      "Get Button Feedback" : "Push Button: State Changes";
   END_VAR
   VAR_TEMP
      feedback : "Push Button Data: State Change Data";
   END_VAR
BEGIN
   REGION "PROCESS USER INPUT"
       #"Get Button Feedback"(interface := #interface,
                              state_changes := #feedback);
   END_REGION

   REGION "ANIMATIONS"

       REGION "COLOR"
           #interface.animate := "Bool.Animate"(true_color := "GREEN_LIGHT_BACKGROUND",
                                                false_color := "GRAY_BACKGROUND",
                                                evaluation_signal := #feedback.actuate.actual);
       END_REGION

       REGION "VISIBILITY"
           #interface.visible := NOT #hide;
       END_REGION

       REGION "ENABLED STATE"
           #interface.enable := NOT #hide;
       END_REGION

   END_REGION

   REGION "SET FIRST ROW"
       IF #feedback.actuate.rising THEN
           #first_row := "NavBar: Private: First Row"(first_row := #first_row,
                                                      offset := -1 * (#VISIBLE_ROW_COUNT + 1),
                                                      TABLE_LENGTH := #TABLE_LENGTH);
       END_IF;
   END_REGION
END_FUNCTION_BLOCK

FUNCTION_BLOCK "NavBar: Page Down"   // FB37, SCL
{ S7_Optimized_Access := 'TRUE' }
VERSION : 0.1
   VAR_INPUT
      hide : Bool;
      TABLE_LENGTH : DInt;
      VISIBLE_ROW_COUNT : DInt;
   END_VAR
   VAR_IN_OUT
      interface : "Push Button Data";
      first_row : DInt;
   END_VAR
   VAR
      "Get Button Feedback" : "Push Button: State Changes";
   END_VAR
   VAR_TEMP
      feedback : "Push Button Data: State Change Data";
   END_VAR
BEGIN
   REGION "PROCESS USER INPUT"
       #"Get Button Feedback"(interface := #interface,
                              state_changes := #feedback);
   END_REGION

   REGION "ANIMATIONS"

       REGION "COLOR"
           #interface.animate := "Bool.Animate"(true_color := "GREEN_LIGHT_BACKGROUND",
                                                false_color := "GRAY_BACKGROUND",
                                                evaluation_signal := #feedback.actuate.actual);
       END_REGION

       REGION "VISIBILITY"
           #interface.visible := NOT #hide;
       END_REGION

       REGION "ENABLED STATE"
           #interface.enable := NOT #hide;
       END_REGION

   END_REGION

   REGION "SET FIRST ROW"
       IF #feedback.actuate.rising THEN
           #first_row := "NavBar: Private: First Row"(first_row := #first_row,
                                                      offset := #VISIBLE_ROW_COUNT + 1,
                                                      TABLE_LENGTH := #TABLE_LENGTH);
       END_IF;
   END_REGION
END_FUNCTION_BLOCK

FUNCTION_BLOCK "NavBar: Line Down"   // FB38, SCL
{ S7_Optimized_Access := 'TRUE' }
VERSION : 0.1
   VAR_INPUT
      hide : Bool;
      TABLE_LENGTH : DInt;
   END_VAR
   VAR_IN_OUT
      interface : "Push Button Data";
      first_row : DInt;
   END_VAR
   VAR
      "Get Button Feedback" : "Push Button: State Changes";
   END_VAR
   VAR_TEMP
      feedback : "Push Button Data: State Change Data";
   END_VAR
BEGIN
   REGION "PROCESS USER INPUT"
       #"Get Button Feedback"(interface := #interface,
                              state_changes := #feedback);
   END_REGION

   REGION "ANIMATIONS"

       REGION "COLOR"
           #interface.animate := "Bool.Animate"(true_color := "GREEN_LIGHT_BACKGROUND",
                                                false_color := "GRAY_BACKGROUND",
                                                evaluation_signal := #feedback.actuate.actual);
       END_REGION

       REGION "VISIBILITY"
           #interface.visible := NOT #hide;
       END_REGION

       REGION "ENABLED STATE"
           #interface.enable := NOT #hide;
       END_REGION

   END_REGION

   REGION "SET FIRST ROW"
       IF #feedback.actuate.rising THEN
           #first_row := "NavBar: Private: First Row"(first_row := #first_row,
                                                      offset := 1,
                                                      TABLE_LENGTH := #TABLE_LENGTH);
       END_IF;
   END_REGION
END_FUNCTION_BLOCK

FUNCTION_BLOCK "NavBar: Line Up"   // FB39, SCL
{ S7_Optimized_Access := 'TRUE' }
VERSION : 0.1
   VAR_INPUT
      hide : Bool;
      TABLE_LENGTH : DInt;
   END_VAR
   VAR_IN_OUT
      interface : "Push Button Data";
      first_row : DInt;
   END_VAR
   VAR
      "Get Button Feedback" : "Push Button: State Changes";
   END_VAR
   VAR_TEMP
      feedback : "Push Button Data: State Change Data";
   END_VAR
BEGIN
   REGION "PROCESS USER INPUT"
       #"Get Button Feedback"(interface := #interface,
                              state_changes := #feedback);
   END_REGION

   REGION "ANIMATIONS"

       REGION "COLOR"
           #interface.animate := "Bool.Animate"(true_color := "GREEN_LIGHT_BACKGROUND",
                                                false_color := "GRAY_BACKGROUND",
                                                evaluation_signal := #feedback.actuate.actual);
       END_REGION

       REGION "VISIBILITY"
           #interface.visible := NOT #hide;
       END_REGION

       REGION "ENABLED STATE"
           #interface.enable := NOT #hide;
       END_REGION

   END_REGION

   REGION "SET FIRST ROW"
       IF #feedback.actuate.rising THEN
           #first_row := "NavBar: Private: First Row"(first_row := #first_row,
                                                      offset := -1,
                                                      TABLE_LENGTH := #TABLE_LENGTH);
       END_IF;
   END_REGION
END_FUNCTION_BLOCK

FUNCTION_BLOCK "NavBar"   // FB40, SCL
{ S7_Optimized_Access := 'TRUE' }
VERSION : 0.1
   VAR_INPUT
      hide : Bool;
      TABLE_LENGTH : DInt := 49;
      VISIBLE_ROW_COUNT : DInt := 2;
   END_VAR
   VAR_IN_OUT
      interface : "Nav Bar Data";
      first_row : DInt;
   END_VAR
   VAR
      Top : "NavBar: Top";
      "Page Up" : "NavBar: Page Up";
      "Line Up" : "NavBar: Line Up";
      "Line Down" : "NavBar: Line Down";
      "Page Down" : "NavBar: Page Down";
      Bottom : "NavBar: Bottom";
   END_VAR
BEGIN
   REGION "BUFFER IN"
       "NavBar: Map HMI to PLC"(hmi := #interface.hmi,
                                plc := #interface.plc);
   END_REGION

   REGION "NAVBAR TOP "
       #Top(hide := #hide,
            TABLE_LENGTH := #TABLE_LENGTH,
            interface := #interface.plc.top,
            first_row := #first_row);
   END_REGION

   REGION "PAGE UP"
       #"Page Up"(hide := #hide,
                  TABLE_LENGTH := #TABLE_LENGTH,
                  VISIBLE_ROW_COUNT := #VISIBLE_ROW_COUNT,
                  interface := #interface.plc.pageUp,
                  first_row := #first_row);
   END_REGION

   REGION "LINE UP"
       #"Line Up"(hide := #hide,
                  TABLE_LENGTH := #TABLE_LENGTH,
                  interface := #interface.plc.lineUp,
                  first_row := #first_row);
   END_REGION

   REGION "LINE DOWN"
       #"Line Down"(hide := #hide,
                    TABLE_LENGTH := #TABLE_LENGTH,
                    interface := #interface.plc.lineDown,
                    first_row := #first_row);
   END_REGION

   REGION "PAGE DOWN"
       #"Page Down"(hide := #hide,
                    TABLE_LENGTH := #TABLE_LENGTH,
                    VISIBLE_ROW_COUNT := #VISIBLE_ROW_COUNT,
                    interface := #interface.plc.pageDown,
                    first_row := #first_row);
   END_REGION

   REGION "BOTTOM"
       #Bottom(hide := #hide,
               TABLE_LENGTH := #TABLE_LENGTH,
               VISIBLE_ROW_COUNT := #VISIBLE_ROW_COUNT,
               interface := #interface.plc.bottom,
               first_row := #first_row);
   END_REGION

   REGION "BUFFER OUT"
       "NavBar: Map PLC to HMI"(plc := #interface.plc,
                                hmi := #interface.hmi);
   END_REGION
END_FUNCTION_BLOCK

FUNCTION "NavBar: Map HMI to PLC" : Void   // FC98, SCL
{ S7_Optimized_Access := 'TRUE' }
VERSION : 0.1
   VAR_INPUT
      hmi : "Nav Bar Data: HMI";
   END_VAR
   VAR_IN_OUT
      plc : "Nav Bar Data: PLC";
   END_VAR
BEGIN
   REGION "NOTES"
       // mapping is necessary because hmi faceplate data structures
       // cannot consist of embedded udts
   END_REGION


   REGION "TOP"
       #plc.top.actuate := #hmi.top_actuate;
       #plc.top.animate := #hmi.top_animate;
       #plc.top.enable := #hmi.top_enable;
       #plc.top.label := #hmi.top_label;
       #plc.top.listSelect := #hmi.top_list_select;
       #plc.top.visible := #hmi.top_visible;
   END_REGION


   REGION "PAGE UP"
       #plc.pageUp.actuate := #hmi.page_up_actuate;
       #plc.pageUp.animate := #hmi.page_up_animate;
       #plc.pageUp.enable := #hmi.page_up_enable;
       #plc.pageUp.label := #hmi.page_up_label;
       #plc.pageUp.listSelect := #hmi.page_up_list_select;
       #plc.pageUp.visible := #hmi.page_up_visible;
   END_REGION


   REGION "LINE UP"
       #plc.lineUp.actuate := #hmi.line_up_actuate;
       #plc.lineUp.animate := #hmi.line_up_animate;
       #plc.lineUp.enable := #hmi.line_up_enable;
       #plc.lineUp.label := #hmi.line_up_label;
       #plc.lineUp.listSelect := #hmi.line_up_list_select;
       #plc.lineUp.visible := #hmi.line_up_visible;
   END_REGION


   REGION "LINE DOWN"
       #plc.lineDown.actuate := #hmi.line_down_actuate;
       #plc.lineDown.animate := #hmi.line_down_animate;
       #plc.lineDown.enable := #hmi.line_down_enable;
       #plc.lineDown.label := #hmi.line_down_label;
       #plc.lineDown.listSelect := #hmi.line_down_list_select;
       #plc.lineDown.visible := #hmi.line_down_visible;
   END_REGION


   REGION "PAGE DOWN"
       #plc.pageDown.actuate := #hmi.page_down_actuate;
       #plc.pageDown.animate := #hmi.page_down_animate;
       #plc.pageDown.enable := #hmi.page_down_enable;
       #plc.pageDown.label := #hmi.page_down_label;
       #plc.pageDown.listSelect := #hmi.page_down_list_select;
       #plc.pageDown.visible := #hmi.page_down_visible;
   END_REGION


   REGION "BOTTOM"
       #plc.bottom.actuate := #hmi.bottom_actuate;
       #plc.bottom.animate := #hmi.bottom_animate;
       #plc.bottom.enable := #hmi.bottom_enable;
       #plc.bottom.label := #hmi.bottom_label;
       #plc.bottom.listSelect := #hmi.bottom_list_select;
       #plc.bottom.visible := #hmi.bottom_visible;
   END_REGION
END_FUNCTION

FUNCTION "NavBar: Map PLC to HMI" : Void   // FC99, SCL
{ S7_Optimized_Access := 'TRUE' }
VERSION : 0.1
   VAR_INPUT
      plc : "Nav Bar Data: PLC";
   END_VAR
   VAR_IN_OUT
      hmi : "Nav Bar Data: HMI";
   END_VAR
BEGIN
   REGION "NOTES"
       // mapping is necessary because hmi faceplate data structures
       // cannot consist of embedded udts
   END_REGION


   REGION "TOP"
       //#hmi.top_actuate := #plc.top.actuate;
       #hmi.top_animate := #plc.top.animate;
       #hmi.top_enable := #plc.top.enable;
       #hmi.top_label := #plc.top.label;
       #hmi.top_list_select := #plc.top.listSelect;
       #hmi.top_visible := #plc.top.visible;
   END_REGION


